WB2[80].2'; 2563 '~Spare WB2[80].3'; 2564 '~S002TT1 VFD Temperature Warning WB2[80].4'; 2565 '~Spare WB2[80].5'; 2566 '~Spare WB2[80].6'; 2567 '~S002TT1 Fixture A Bypass Selected WB2[80].7'; 2568 '~S002TT1 Fixture B Bypass Selected WB2[80].8'; 2569 '~S002TT1 Fixture C Bypass Selected WB2[80].9'; 2570 '~S002TT1 Fixture D Bypass Selected WB2[80].10'; 2571 '~S002TT1 Fixture E Bypass Selected WB2[80].11'; 2572 '~S002TT1 Fixture F Bypass Selected WB2[80].12'; 2573 '~S002TT1 Manual Mode Motion Not Enabled WB2[80].13'; 2574 '~S002TT1 Lt Screen Not Clear Or Active WB2[80].14'; 2575 '~S002TT1 Robots Not Clear Of Turntable Index WB2[80].15'; 2576 '~S002TT1 All Tooling Not Clear To Rotate WB2[80].16'; 2577 '~S002TT1 Turn Table Brake Still Released WB2[80].17'; 2578 '~S002TT1DES1 - S002TT1 EtherNet Switch Port At Half Duplex WB2[80].18'; 2579 '~S002TT1DES1 - S002TT1 EtherNet Switch Config Changes Not Saved WB2[80].19'; 2580 '~S002TT1DES1 - S002TT1 EtherNet Switch Configuration Changed WB2[80].20'; 2581 '~S002TT1DES1 - S002TT1 EtherNet Switch Port With Excessive Errors WB2[80].21'; 2582 '~S002TT1DES1 - S002TT1 EtherNet Switch Port With Utilization Warn WB2[80].22'; 2583 '~S002TT1DES1 - S002TT1 EtherNet Switch Changes Require Reboot WB2[80].23'; 2584 '~Spare WB2[80].24'; 2585 '~S002TT1DES2 - S002TT1 EtherNet Switch Port At Half Duplex WB2[80].25'; 2586 '~S002TT1DES2 - S002TT1 EtherNet Switch Config Changes Not Saved WB2[80].26'; 2587 '~S002TT1DES2 - S002TT1 EtherNet Switch Configuration Changed WB2[80].27'; 2588 '~S002TT1DES2 - S002TT1 EtherNet Switch Port With Excessive Errors WB2[80].28'; 2589 '~S002TT1DES2 - S002TT1 EtherNet Switch Port With Utilization Warn WB2[80].29'; 2590 '~S002TT1DES2 - S002TT1 EtherNet Switch Changes Require Reboot WB2[80].30'; 2591 '~Spare WB2[80].31'; 2592 '~Spare WB2[81].0'; 2593 '~Spare WB2[81].1'; 2594 '~Spare WB2[81].2'; 2595 '~Spare WB2[81].3'; 2596 '~Spare WB2[81].4'; 2597 '~Spare WB2[81].5'; 2598 '~Spare WB2[81].6'; 2599 '~Spare WB2[81].7'; 2600 '~Spare WB2[81].8'; 2601 '~Spare WB2[81].9'; 2602 '~Spare WB2[81].10'; 2603 '~Spare WB2[81].11'; 2604 '~Spare WB2[81].12'; 2605 '~Spare WB2[81].13'; 2606 '~Spare WB2[81].14'; 2607 '~Spare WB2[81].15'; 2608 '~Spare WB2[81].16'; 2609 '~Spare WB2[81].17'; 2610 '~Spare WB2[81].18'; 2611 '~Spare WB2[81].19'; 2612 '~Spare WB2[81].20'; 2613 '~Spare WB2[81].21'; 2614 '~Spare WB2[81].22'; 2615 '~Spare WB2[81].23'; 2616 '~Spare WB2[81].24'; 2617 '~Spare WB2[81].25'; 2618 '~Spare WB2[81].26'; 2619 '~Spare WB2[81].27'; 2620 '~Spare WB2[81].28'; 2621 '~Spare WB2[81].29'; 2622 '~Spare WB2[81].30'; 2623 '~Spare WB2[81].31'; 2624 '~Spare WB2[82].0'; 2625 '~Spare WB2[82].1'; 2626 '~Spare WB2[82].2'; 2627 '~Spare WB2[82].3'; 2628 '~Spare WB2[82].4'; 2629 '~Spare WB2[82].5'; 2630 '~Spare WB2[82].6'; 2631 '~Spare WB2[82].7'; 2632 '~Spare WB2[82].8'; 2633 '~Spare WB2[82].9'; 2634 '~Spare WB2[82].10'; 2635 '~Spare WB2[82].11'; 2636 '~Spare WB2[82].12'; 2637 '~Spare WB2[82].13'; 2638 '~Spare WB2[82].14'; 2639 '~Spare WB2[82].15'; 2640 '~Spare WB2[82].16'; 2641 '~Spare WB2[82].17'; 2642 '~Spare WB2[82].18'; 2643 '~Spare WB2[82].19'; 2644 '~Spare WB2[82].20'; 2645 '~Spare WB2[82].21'; 2646 '~Spare WB2[82].22'; 2647 '~Spare WB2[82].23'; 2648 '~Spare WB2[82].24'; 2649 '~Spare WB2[82].25'; 2650 '~Spare WB2[82].26'; 2651 '~Spare WB2[82].27'; 2652 '~Spare WB2[82].28'; 2653 '~Spare WB2[82].29'; 2654 '~Spare WB2[82].30'; 2655 '~Spare WB2[82].31'; 2656 '~Spare WB2[83].0'; 2657 '~Spare WB2[83].1'; 2658 '~Spare WB2[83].2'; 2659 '~Spare WB2[83].3'; 2660 '~Spare WB2[83].4'; 2661 '~Spare WB2[83].5'; 2662 '~Spare WB2[83].6'; 2663 '~Spare WB2[83].7'; 2664 '~Spare WB2[83].8'; 2665 '~Spare WB2[83].9'; 2666 '~Spare WB2[83].10'; 2667 '~Spare WB2[83].11'; 2668 '~Spare WB2[83].12'; 2669 '~Spare WB2[83].13'; 2670 '~Spare WB2[83].14'; 2671 '~Spare WB2[83].15'; 2672 '~Spare WB2[83].16'; 2673 '~Spare WB2[83].17'; 2674 '~Spare WB2[83].18'; 2675 '~Spare WB2[83].19'; 2676 '~Spare WB2[83].20'; 2677 '~Spare WB2[83].21'; 2678 '~Spare WB2[83].22'; 2679 '~Spare WB2[83].23'; 2680 '~Spare WB2[83].24'; 2681 '~Spare WB2[83].25'; 2682 '~Spare WB2[83].26'; 2683 '~Spare WB2[83].27'; 2684 '~Spare WB2[83].28'; 2685 '~Spare WB2[83].29'; 2686 '~Spare WB2[83].30'; 2687 '~Spare WB2[83].31'; 2688 '~S001PRB Overtime WB2[84].0'; 2689 '~S001PRB - VFD Temperature Warning WB2[84].1'; 2690 '~Spare WB2[84].2'; 2691 '~S001PRB Coded Rail Reader Optics Alarm WB2[84].3'; 2692 '~S001PRB Coded Rail Reader Data Not Valid WB2[84].4'; 2693 '~S001PRB Brake Still Released WB2[84].5'; 2694 '~Spare WB2[84].6'; 2695 '~S001LFT Brake Still Released WB2[84].7'; 2696 '~S001PRB - PRB VFD Heatsink Fan Should Be Replaced WB2[84].8'; 2697 '~S001PRB - PRB VFD Internal Fan Should Be Replaced WB2[84].9'; 2698 '~S002PRB Overtime WB2[84].10'; 2699 '~S002PRB - VFD Temperature Warning WB2[84].11'; 2700 '~Spare WB2[84].12'; 2701 '~S002PRB Coded Rail Reader Optics Alarm WB2[84].13'; 2702 '~S002PRB Coded Rail Reader Data Not Valid WB2[84].14'; 2703 '~S002PRB Brake Still Released WB2[84].15'; 2704 '~Spare WB2[84].16'; 2705 '~S002LFT Brake Still Released WB2[84].17'; 2706 '~S002PRB - PRB VFD Heatsink Fan Should Be Replaced WB2[84].18'; 2707 '~S002PRB - PRB VFD Internal Fan Should Be Replaced WB2[84].19'; 2708 '~Spare WB2[84].20'; 2709 '~Spare WB2[84].21'; 2710 '~Spare WB2[84].22'; 2711 '~Spare WB2[84].23'; 2712 '~Spare WB2[84].24'; 2713 '~S001_002PRBDES1 - EtherNet Switch Port At Half Duplex WB2[84].25'; 2714 '~S001_002PRBDES1 - EtherNet Switch Configuration Changes Not Saved WB2[84].26'; 2715 '~S001_002PRBDES1 - EtherNet Switch Configuration Changed WB2[84].27'; 2716 '~S001_002PRBDES1 - EtherNet Switch Port With Excessive Errors WB2[84].28'; 2717 '~S001_002PRBDES1 - EtherNet Switch Port With Utilization Warning WB2[84].29'; 2718 '~S001_002PRBDES1 - EtherNet Switch Changes Require Reboot WB2[84].30'; 2719 '~Spare WB2[84].31'; 2720 '~S003PRB Overtime WB2[85].0'; 2721 '~S003PRB VFD Temperature Warning WB2[85].1'; 2722 '~Spare WB2[85].2'; 2723 '~Spare WB2[85].3'; 2724 '~Spare WB2[85].4'; 2725 '~S003PRB Brake Still Released WB2[85].5'; 2726 '~S003PRB Running Low Speed In Auto WB2[85].6'; 2727 '~S003LFT Brake Still Released WB2[85].7'; 2728 '~Spare WB2[85].8'; 2729 '~Spare WB2[85].9'; 2730 '~S004PRB Overtime WB2[85].10'; 2731 '~S004PRB VFD Temperature Warning WB2[85].11'; 2732 '~Spare WB2[85].12'; 2733 '~Spare WB2[85].13'; 2734 '~Spare WB2[85].14'; 2735 '~S004PRB Brake Still Released WB2[85].15'; 2736 '~S004PRB Running Low Speed In Auto WB2[85].16'; 2737 '~S004LFT Brake Still Released WB2[85].17'; 2738 '~Spare WB2[85].18'; 2739 '~Spare WB2[85].19'; 2740 '~Spare WB2[85].20'; 2741 '~Spare WB2[85].21'; 2742 '~Spare WB2[85].22'; 2743 '~Spare WB2[85].23'; 2744 '~Spare WB2[85].24'; 2745 '~S003_004PRBDES1 - EtherNet Switch Port At Half Duplex WB2[85].25'; 2746 '~S003_004PRBDES1 - EtherNet Switch Configuration Changes Not Saved WB2[85].26'; 2747 '~S003_004PRBDES1 - EtherNet Switch Configuration Changed WB2[85].27'; 2748 '~S003_004PRBDES1 - EtherNet Switch Port With Excessive Errors WB2[85].28'; 2749 '~S003_004PRBDES1 - EtherNet Switch Port With Utilization Warning WB2[85].29'; 2750 '~S003_004PRBDES1 - EtherNet Switch Changes Require Reboot WB2[85].30'; 2751 '~Spare WB2[85].31'; 2752 '~Spare WB2[86].0'; 2753 '~Spare WB2[86].1'; 2754 '~Spare WB2[86].2'; 2755 '~Spare WB2[86].3'; 2756 '~Spare WB2[86].4'; 2757 '~Spare WB2[86].5'; 2758 '~Spare WB2[86].6'; 2759 '~Spare WB2[86].7'; 2760 '~Spare WB2[86].8'; 2761 '~Spare WB2[86].9'; 2762 '~Spare WB2[86].10'; 2763 '~Spare WB2[86].11'; 2764 '~Spare WB2[86].12'; 2765 '~Spare WB2[86].13'; 2766 '~Spare WB2[86].14'; 2767 '~Spare WB2[86].15'; 2768 '~Spare WB2[86].16'; 2769 '~Spare WB2[86].17'; 2770 '~Spare WB2[86].18'; 2771 '~Spare WB2[86].19'; 2772 '~Spare WB2[86].20'; 2773 '~Spare WB2[86].21'; 2774 '~Spare WB2[86].22'; 2775 '~Spare WB2[86].23'; 2776 '~Spare WB2[86].24'; 2777 '~Spare WB2[86].25'; 2778 '~Spare WB2[86].26'; 2779 '~Spare WB2[86].27'; 2780 '~Spare WB2[86].28'; 2781 '~Spare WB2[86].29'; 2782 '~Spare WB2[86].30'; 2783 '~Spare WB2[86].31'; 2784 '~Spare WB2[87].0'; 2785 '~Spare WB2[87].1'; 2786 '~Spare WB2[87].2'; 2787 '~Spare WB2[87].3'; 2788 '~Spare WB2[87].4'; 2789 '~Spare WB2[87].5'; 2790 '~Spare WB2[87].6'; 2791 '~Spare WB2[87].7'; 2792 '~Spare WB2[87].8'; 2793 '~Spare WB2[87].9'; 2794 '~Spare WB2[87].10'; 2795 '~Spare WB2[87].11'; 2796 '~Spare WB2[87].12'; 2797 '~Spare WB2[87].13'; 2798 '~Spare WB2[87].14'; 2799 '~Spare WB2[87].15'; 2800 '~Spare WB2[87].16'; 2801 '~Spare WB2[87].17'; 2802 '~Spare WB2[87].18'; 2803 '~Spare WB2[87].19'; 2804 '~Spare WB2[87].20'; 2805 '~Spare WB2[87].21'; 2806 '~Spare WB2[87].22'; 2807 '~Spare WB2[87].23'; 2808 '~Spare WB2[87].24'; 2809 '~Spare WB2[87].25'; 2810 '~Spare WB2[87].26'; 2811 '~Spare WB2[87].27'; 2812 '~Spare WB2[87].28'; 2813 '~Spare WB2[87].29'; 2814 '~Spare WB2[87].30'; 2815 '~Spare WB2[87].31'; 2816 '~Spare WB2[88].0'; 2817 '~Spare WB2[88].1'; 2818 '~Spare WB2[88].2'; 2819 '~Spare WB2[88].3'; 2820 '~Spare WB2[88].4'; 2821 '~Spare WB2[88].5'; 2822 '~Spare WB2[88].6'; 2823 '~Spare WB2[88].7'; 2824 '~Spare WB2[88].8'; 2825 '~Spare WB2[88].9'; 2826 '~Spare WB2[88].10'; 2827 '~Spare WB2[88].11'; 2828 '~Spare WB2[88].12'; 2829 '~Spare WB2[88].13'; 2830 '~Spare WB2[88].14'; 2831 '~Spare WB2[88].15'; 2832 '~Spare WB2[88].16'; 2833 '~Spare WB2[88].17'; 2834 '~Spare WB2[88].18'; 2835 '~Spare WB2[88].19'; 2836 '~Spare WB2[88].20'; 2837 '~Spare WB2[88].21'; 2838 '~Spare WB2[88].22'; 2839 '~Spare WB2[88].23'; 2840 '~Spare WB2[88].24'; 2841 '~Spare WB2[88].25'; 2842 '~Spare WB2[88].26'; 2843 '~Spare WB2[88].27'; 2844 '~Spare WB2[88].28'; 2845 '~Spare WB2[88].29'; 2846 '~Spare WB2[88].30'; 2847 '~Spare WB2[88].31'; 2848 '~Spare WB2[89].0'; 2849 '~Spare WB2[89].1'; 2850 '~Spare WB2[89].2'; 2851 '~Spare WB2[89].3'; 2852 '~Spare WB2[89].4'; 2853 '~Spare WB2[89].5'; 2854 '~Spare WB2[89].6'; 2855 '~Spare WB2[89].7'; 2856 '~Spare WB2[89].8'; 2857 '~Spare WB2[89].9'; 2858 '~Spare WB2[89].10'; 2859 '~Spare WB2[89].11'; 2860 '~Spare WB2[89].12'; 2861 '~Spare WB2[89].13'; 2862 '~Spare WB2[89].14'; 2863 '~Spare WB2[89].15'; 2864 '~Spare WB2[89].16'; 2865 '~Spare WB2[89].17'; 2866 '~Spare WB2[89].18'; 2867 '~Spare WB2[89].19'; 2868 '~Spare WB2[89].20'; 2869 '~Spare WB2[89].21'; 2870 '~Spare WB2[89].22'; 2871 '~Spare WB2[89].23'; 2872 '~Spare WB2[89].24'; 2873 '~Spare WB2[89].25'; 2874 '~Spare WB2[89].26'; 2875 '~Spare WB2[89].27'; 2876 '~Spare WB2[89].28'; 2877 '~Spare WB2[89].29'; 2878 '~Spare WB2[89].30'; 2879 '~Spare WB2[89].31'; 2880 '~Spare WB2[90].0'; 2881 '~Spare WB2[90].1'; 2882 '~Spare WB2[90].2'; 2883 '~Spare WB2[90].3'; 2884 '~Spare WB2[90].4'; 2885 '~Spare WB2[90].5'; 2886 '~Spare WB2[90].6'; 2887 '~Spare WB2[90].7'; 2888 '~Spare WB2[90].8'; 2889 '~Spare WB2[90].9'; 2890 '~Spare WB2[90].10'; 2891 '~Spare WB2[90].11'; 2892 '~Spare WB2[90].12'; 2893 '~Spare WB2[90].13'; 2894 '~Spare WB2[90].14'; 2895 '~Spare WB2[90].15'; 2896 '~Spare WB2[90].16'; 2897 '~Spare WB2[90].17'; 2898 '~Spare WB2[90].18'; 2899 '~Spare WB2[90].19'; 2900 '~Spare WB2[90].20'; 2901 '~Spare WB2[90].21'; 2902 '~Spare WB2[90].22'; 2903 '~Spare WB2[90].23'; 2904 '~Spare WB2[90].24'; 2905 '~Spare WB2[90].25'; 2906 '~Spare WB2[90].26'; 2907 '~Spare WB2[90].27'; 2908 '~Spare WB2[90].28'; 2909 '~Spare WB2[90].29'; 2910 '~Spare WB2[90].30'; 2911 '~Spare WB2[90].31'; 2912 '~Spare WB2[91].0'; 2913 '~Spare WB2[91].1'; 2914 '~Spare WB2[91].2'; 2915 '~Spare WB2[91].3'; 2916 '~Spare WB2[91].4'; 2917 '~Spare WB2[91].5'; 2918 '~Spare WB2[91].6'; 2919 '~Spare WB2[91].7'; 2920 '~Spare WB2[91].8'; 2921 '~Spare WB2[91].9'; 2922 '~Spare WB2[91].10'; 2923 '~Spare WB2[91].11'; 2924 '~Spare WB2[91].12'; 2925 '~Spare WB2[91].13'; 2926 '~Spare WB2[91].14'; 2927 '~Spare WB2[91].15'; 2928 '~Spare WB2[91].16'; 2929 '~Spare WB2[91].17'; 2930 '~Spare WB2[91].18'; 2931 '~Spare WB2[91].19'; 2932 '~Spare WB2[91].20'; 2933 '~Spare WB2[91].21'; 2934 '~Spare WB2[91].22'; 2935 '~Spare WB2[91].23'; 2936 '~Spare WB2[91].24'; 2937 '~Spare WB2[91].25'; 2938 '~Spare WB2[91].26'; 2939 '~Spare WB2[91].27'; 2940 '~Spare WB2[91].28'; 2941 '~Spare WB2[91].29'; 2942 '~Spare WB2[91].30'; 2943 '~Spare WB2[91].31'; 2944 '~Spare WB2[92].0'; 2945 '~Spare WB2[92].1'; 2946 '~Spare WB2[92].2'; 2947 '~Spare WB2[92].3'; 2948 '~Spare WB2[92].4'; 2949 '~Spare WB2[92].5'; 2950 '~Spare WB2[92].6'; 2951 '~Spare WB2[92].7'; 2952 '~Spare WB2[92].8'; 2953 '~Spare WB2[92].9'; 2954 '~Spare WB2[92].10'; 2955 '~Spare WB2[92].11'; 2956 '~Spare WB2[92].12'; 2957 '~Spare WB2[92].13'; 2958 '~Spare WB2[92].14'; 2959 '~Spare WB2[92].15'; 2960 '~Spare WB2[92].16'; 2961 '~Spare WB2[92].17'; 2962 '~Spare WB2[92].18'; 2963 '~Spare WB2[92].19'; 2964 '~Spare WB2[92].20'; 2965 '~Spare WB2[92].21'; 2966 '~Spare WB2[92].22'; 2967 '~Spare WB2[92].23'; 2968 '~Spare WB2[92].24'; 2969 '~Spare WB2[92].25'; 2970 '~Spare WB2[92].26'; 2971 '~Spare WB2[92].27'; 2972 '~Spare WB2[92].28'; 2973 '~Spare WB2[92].29'; 2974 '~Spare WB2[92].30'; 2975 '~Spare WB2[92].31'; 2976 '~Spare WB2[93].0'; 2977 '~Spare WB2[93].1'; 2978 '~Spare WB2[93].2'; 2979 '~Spare WB2[93].3'; 2980 '~Spare WB2[93].4'; 2981 '~Spare WB2[93].5'; 2982 '~Spare WB2[93].6'; 2983 '~Spare WB2[93].7'; 2984 '~Spare WB2[93].8'; 2985 '~Spare WB2[93].9'; 2986 '~Spare WB2[93].10'; 2987 '~Spare WB2[93].11'; 2988 '~Spare WB2[93].12'; 2989 '~Spare WB2[93].13'; 2990 '~Spare WB2[93].14'; 2991 '~Spare WB2[93].15'; 2992 '~Spare WB2[93].16'; 2993 '~Spare WB2[93].17'; 2994 '~Spare WB2[93].18'; 2995 '~Spare WB2[93].19'; 2996 '~Spare WB2[93].20'; 2997 '~Spare WB2[93].21'; 2998 '~Spare WB2[93].22'; 2999 '~Spare WB2[93].23'; 3000 '~Spare WB2[93].24'; 3001 '~Spare WB2[93].25'; 3002 '~Spare WB2[93].26'; 3003 '~Spare WB2[93].27'; 3004 '~Spare WB2[93].28'; 3005 '~Spare WB2[93].29'; 3006 '~Spare WB2[93].30'; 3007 '~Spare WB2[93].31'; 3008 '~Spare WB2[94].0'; 3009 '~Spare WB2[94].1'; 3010 '~Spare WB2[94].2'; 3011 '~Spare WB2[94].3'; 3012 '~Spare WB2[94].4'; 3013 '~Spare WB2[94].5'; 3014 '~Spare WB2[94].6'; 3015 '~Spare WB2[94].7'; 3016 '~Spare WB2[94].8'; 3017 '~Spare WB2[94].9'; 3018 '~Spare WB2[94].10'; 3019 '~Spare WB2[94].11'; 3020 '~Spare WB2[94].12'; 3021 '~Spare WB2[94].13'; 3022 '~Spare WB2[94].14'; 3023 '~Spare WB2[94].15'; 3024 '~Spare WB2[94].16'; 3025 '~Spare WB2[94].17'; 3026 '~Spare WB2[94].18'; 3027 '~Spare WB2[94].19'; 3028 '~Spare WB2[94].20'; 3029 '~Spare WB2[94].21'; 3030 '~Spare WB2[94].22'; 3031 '~Spare WB2[94].23'; 3032 '~Spare WB2[94].24'; 3033 '~Spare WB2[94].25'; 3034 '~Spare WB2[94].26'; 3035 '~Spare WB2[94].27'; 3036 '~Spare WB2[94].28'; 3037 '~Spare WB2[94].29'; 3038 '~Spare WB2[94].30'; 3039 '~Spare WB2[94].31'; 3040 '~Spare WB2[95].0'; 3041 '~Spare WB2[95].1'; 3042 '~Spare WB2[95].2'; 3043 '~Spare WB2[95].3'; 3044 '~Spare WB2[95].4'; 3045 '~Spare WB2[95].5'; 3046 '~Spare WB2[95].6'; 3047 '~Spare WB2[95].7'; 3048 '~Spare WB2[95].8'; 3049 '~Spare WB2[95].9'; 3050 '~Spare WB2[95].10'; 3051 '~Spare WB2[95].11'; 3052 '~Spare WB2[95].12'; 3053 '~Spare WB2[95].13'; 3054 '~Spare WB2[95].14'; 3055 '~Spare WB2[95].15'; 3056 '~Spare WB2[95].16'; 3057 '~Spare WB2[95].17'; 3058 '~Spare WB2[95].18'; 3059 '~Spare WB2[95].19'; 3060 '~Spare WB2[95].20'; 3061 '~Spare WB2[95].21'; 3062 '~Spare WB2[95].22'; 3063 '~Spare WB2[95].23'; 3064 '~Spare WB2[95].24'; 3065 '~Spare WB2[95].25'; 3066 '~Spare WB2[95].26'; 3067 '~Spare WB2[95].27'; 3068 '~Spare WB2[95].28'; 3069 '~Spare WB2[95].29'; 3070 '~Spare WB2[95].30'; 3071 '~Spare WB2[95].31'; 3072 '~Spare WB2[96].0'; 3073 '~Spare WB2[96].1'; 3074 '~Spare WB2[96].2'; 3075 '~Spare WB2[96].3'; 3076 '~Spare WB2[96].4'; 3077 '~Spare WB2[96].5'; 3078 '~Spare WB2[96].6'; 3079 '~Spare WB2[96].7'; 3080 '~Spare WB2[96].8'; 3081 '~Spare WB2[96].9'; 3082 '~Spare WB2[96].10'; 3083 '~Spare WB2[96].11'; 3084 '~Spare WB2[96].12'; 3085 '~Spare WB2[96].13'; 3086 '~Spare WB2[96].14'; 3087 '~Spare WB2[96].15'; 3088 '~Spare WB2[96].16'; 3089 '~Spare WB2[96].17'; 3090 '~Spare WB2[96].18'; 3091 '~Spare WB2[96].19'; 3092 '~Spare WB2[96].20'; 3093 '~Spare WB2[96].21'; 3094 '~Spare WB2[96].22'; 3095 '~Spare WB2[96].23'; 3096 '~Spare WB2[96].24'; 3097 '~Spare WB2[96].25'; 3098 '~Spare WB2[96].26'; 3099 '~Spare WB2[96].27'; 3100 '~Spare WB2[96].28'; 3101 '~Spare WB2[96].29'; 3102 '~Spare WB2[96].30'; 3103 '~Spare WB2[96].31'; 3104 '~Spare WB2[97].0'; 3105 '~Spare WB2[97].1'; 3106 '~Spare WB2[97].2'; 3107 '~Spare WB2[97].3'; 3108 '~Spare WB2[97].4'; 3109 '~Spare WB2[97].5'; 3110 '~Spare WB2[97].6'; 3111 '~Spare WB2[97].7'; 3112 '~Spare WB2[97].8'; 3113 '~Spare WB2[97].9'; 3114 '~Spare WB2[97].10'; 3115 '~Spare WB2[97].11'; 3116 '~Spare WB2[97].12'; 3117 '~Spare WB2[97].13'; 3118 '~Spare WB2[97].14'; 3119 '~Spare WB2[97].15'; 3120 '~Spare WB2[97].16'; 3121 '~Spare WB2[97].17'; 3122 '~Spare WB2[97].18'; 3123 '~Spare WB2[97].19'; 3124 '~Spare WB2[97].20'; 3125 '~Spare WB2[97].21'; 3126 '~Spare WB2[97].22'; 3127 '~Spare WB2[97].23'; 3128 '~Spare WB2[97].24'; 3129 '~Spare WB2[97].25'; 3130 '~Spare WB2[97].26'; 3131 '~Spare WB2[97].27'; 3132 '~Spare WB2[97].28'; 3133 '~Spare WB2[97].29'; 3134 '~Spare WB2[97].30'; 3135 '~Spare WB2[97].31'; 3136 '~Spare WB2[98].0'; 3137 '~Spare WB2[98].1'; 3138 '~Spare WB2[98].2'; 3139 '~Spare WB2[98].3'; 3140 '~Spare WB2[98].4'; 3141 '~Spare WB2[98].5'; 3142 '~Spare WB2[98].6'; 3143 '~Spare WB2[98].7'; 3144 '~Spare WB2[98].8'; 3145 '~Spare WB2[98].9'; 3146 '~Spare WB2[98].10'; 3147 '~Spare WB2[98].11'; 3148 '~Spare WB2[98].12'; 3149 '~Spare WB2[98].13'; 3150 '~Spare WB2[98].14'; 3151 '~Spare WB2[98].15'; 3152 '~Spare WB2[98].16'; 3153 '~Spare WB2[98].17'; 3154 '~Spare WB2[98].18'; 3155 '~Spare WB2[98].19'; 3156 '~Spare WB2[98].20'; 3157 '~Spare WB2[98].21'; 3158 '~Spare WB2[98].22'; 3159 '~Spare WB2[98].23'; 3160 '~Spare WB2[98].24'; 3161 '~Spare WB2[98].25'; 3162 '~Spare WB2[98].26'; 3163 '~Spare WB2[98].27'; 3164 '~Spare WB2[98].28'; 3165 '~Spare WB2[98].29'; 3166 '~Spare WB2[98].30'; 3167 '~Spare WB2[98].31'; 3168 '~Spare WB2[99].0'; 3169 '~Spare WB2[99].1'; 3170 '~Spare WB2[99].2'; 3171 '~Spare WB2[99].3'; 3172 '~Spare WB2[99].4'; 3173 '~Spare WB2[99].5'; 3174 '~Spare WB2[99].6'; 3175 '~Spare WB2[99].7'; 3176 '~Spare WB2[99].8'; 3177 '~Spare WB2[99].9'; 3178 '~Spare WB2[99].10'; 3179 '~Spare WB2[99].11'; 3180 '~Spare WB2[99].12'; 3181 '~Spare WB2[99].13'; 3182 '~Spare WB2[99].14'; 3183 '~Spare WB2[99].15'; 3184 '~Spare WB2[99].16'; 3185 '~Spare WB2[99].17'; 3186 '~Spare WB2[99].18'; 3187 '~Spare WB2[99].19'; 3188 '~Spare WB2[99].20'; 3189 '~Spare WB2[99].21'; 3190 '~Spare WB2[99].22'; 3191 '~Spare WB2[99].23'; 3192 '~Spare WB2[99].24'; 3193 '~Spare WB2[99].25'; 3194 '~Spare WB2[99].26'; 3195 '~Spare WB2[99].27'; 3196 '~Spare WB2[99].28'; 3197 '~Spare WB2[99].29'; 3198 '~Spare WB2[99].30'; 3199 '~S002 Last Message WB2[99].31'

text list "Banner_Scroll Faults": 0 'SCROLL FAULTS ENABLED'; 1 'SCROLL FAULTS DISABLED'

text list "Banner_ScreenName": 1 'Selection Screen'; 3 'Safety Fault'; 19 'PullOff Cart'; 65 'Index Conveyor'; 66 'Belt Conveyor'; 71 'Tip Status1'; 72 'Tip Status2'; 73 'Mig Weld Status1'; 74 'Mig Weld Status2'; 81 'Fixture1 Fault'; 90 'Weld'; 91 'Stepper Reset'; 92 'Rivet'; 100 'Safety N/w. Overview'; 102 'Safety I/O Overview'; 103 'Safety Inst. Overview'; 105 'Safety Inst. Status'; 108 'Enet Network Select'; 109 'Enet Diagnostics'; 1000 'System Screen'; 1001 'User Administration'

